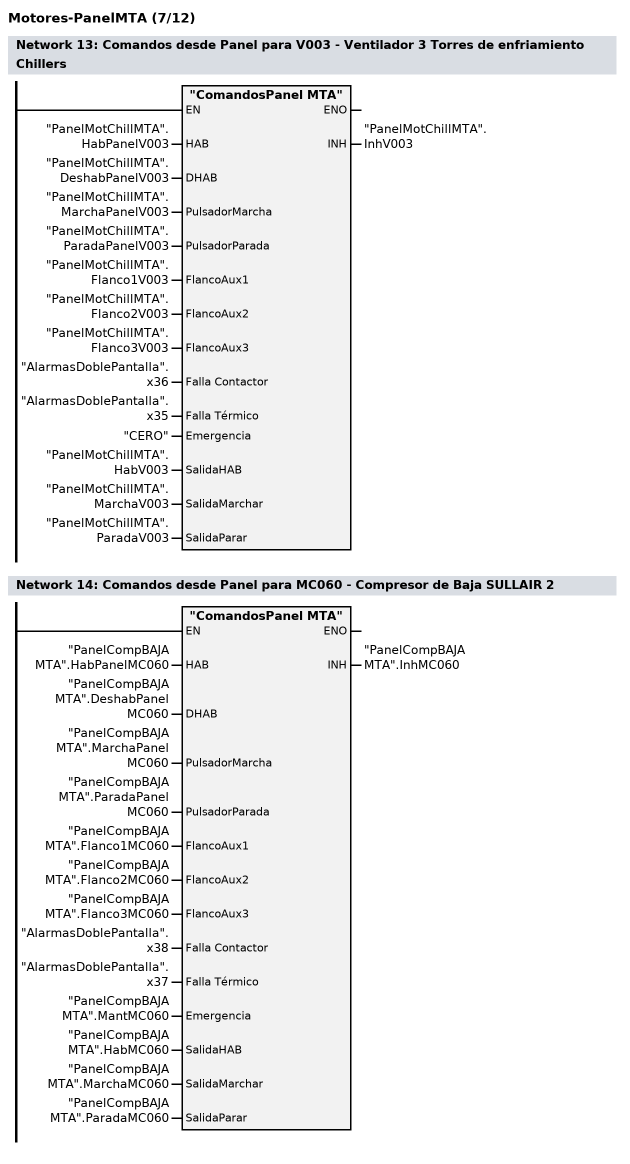
   RUNG wire#powerrail
      "ComandosPanel MTA"(HAB := "PanelMotChillMTA".HabPanelV003, DHAB := "PanelMotChillMTA".DeshabPanelV003, PulsadorMarcha := "PanelMotChillMTA".MarchaPanelV003, PulsadorParada := "PanelMotChillMTA".ParadaPanelV003, FlancoAux1 := "PanelMotChillMTA".Flanco1V003, FlancoAux2 := "PanelMotChillMTA".Flanco2V003, FlancoAux3 := "PanelMotChillMTA".Flanco3V003, "Falla Contactor" := "AlarmasDoblePantalla".x36, "Falla Térmico" := "AlarmasDoblePantalla".x35, Emergencia := "CERO", SalidaHAB := "PanelMotChillMTA".HabV003, SalidaMarchar := "PanelMotChillMTA".MarchaV003, SalidaParar := "PanelMotChillMTA".ParadaV003, INH => "PanelMotChillMTA".InhV003)
   END_RUNG
   // the same network as SCL:
   "ComandosPanel MTA"(HAB := "PanelMotChillMTA".HabPanelV003,
                       DHAB := "PanelMotChillMTA".DeshabPanelV003,
                       PulsadorMarcha := "PanelMotChillMTA".MarchaPanelV003,
                       PulsadorParada := "PanelMotChillMTA".ParadaPanelV003,
                       FlancoAux1 := "PanelMotChillMTA".Flanco1V003,
                       FlancoAux2 := "PanelMotChillMTA".Flanco2V003,
                       FlancoAux3 := "PanelMotChillMTA".Flanco3V003,
                       "Falla Contactor" := "AlarmasDoblePantalla".x36,
                       "Falla Térmico" := "AlarmasDoblePantalla".x35,
                       Emergencia := "CERO",
                       SalidaHAB := "PanelMotChillMTA".HabV003,
                       SalidaMarchar := "PanelMotChillMTA".MarchaV003,
                       SalidaParar := "PanelMotChillMTA".ParadaV003,
                       INH => "PanelMotChillMTA".InhV003);
END_REGION

REGION Network 14: Comandos desde Panel para MC060 - Compresor de Baja SULLAIR 2
   RUNG wire#powerrail
      "ComandosPanel MTA"(HAB := "PanelCompBAJA MTA".HabPanelMC060, DHAB := "PanelCompBAJA MTA".DeshabPanelMC060, PulsadorMarcha := "PanelCompBAJA MTA".MarchaPanelMC060, PulsadorParada := "PanelCompBAJA MTA".ParadaPanelMC060, FlancoAux1 := "PanelCompBAJA MTA".Flanco1MC060, FlancoAux2 := "PanelCompBAJA MTA".Flanco2MC060, FlancoAux3 := "PanelCompBAJA MTA".Flanco3MC060, "Falla Contactor" := "AlarmasDoblePantalla".x38, "Falla Térmico" := "AlarmasDoblePantalla".x37, Emergencia := "PanelCompBAJA MTA".MantMC060, INH => "PanelCompBAJA MTA".InhMC060, SalidaHAB := "PanelCompBAJA MTA".HabMC060, SalidaMarchar := "PanelCompBAJA MTA".MarchaMC060, SalidaParar := "PanelCompBAJA MTA".ParadaMC060)
   END_RUNG
   // the same network as SCL:
   "ComandosPanel MTA"(HAB := "PanelCompBAJA MTA".HabPanelMC060,
                       DHAB := "PanelCompBAJA MTA".DeshabPanelMC060,
                       PulsadorMarcha := "PanelCompBAJA MTA".MarchaPanelMC060,
                       PulsadorParada := "PanelCompBAJA MTA".ParadaPanelMC060,
                       FlancoAux1 := "PanelCompBAJA MTA".Flanco1MC060,
                       FlancoAux2 := "PanelCompBAJA MTA".Flanco2MC060,
                       FlancoAux3 := "PanelCompBAJA MTA".Flanco3MC060,
                       "Falla Contactor" := "AlarmasDoblePantalla".x38,
                       "Falla Térmico" := "AlarmasDoblePantalla".x37,
                       Emergencia := "PanelCompBAJA MTA".MantMC060,
                       SalidaHAB := "PanelCompBAJA MTA".HabMC060,
                       SalidaMarchar := "PanelCompBAJA MTA".MarchaMC060,
                       SalidaParar := "PanelCompBAJA MTA".ParadaMC060,
                       INH => "PanelCompBAJA MTA".InhMC060);
END_REGION

REGION Network 15: Comandos desde Panel para MC061 - Compresor de Baja SULLAIR 1
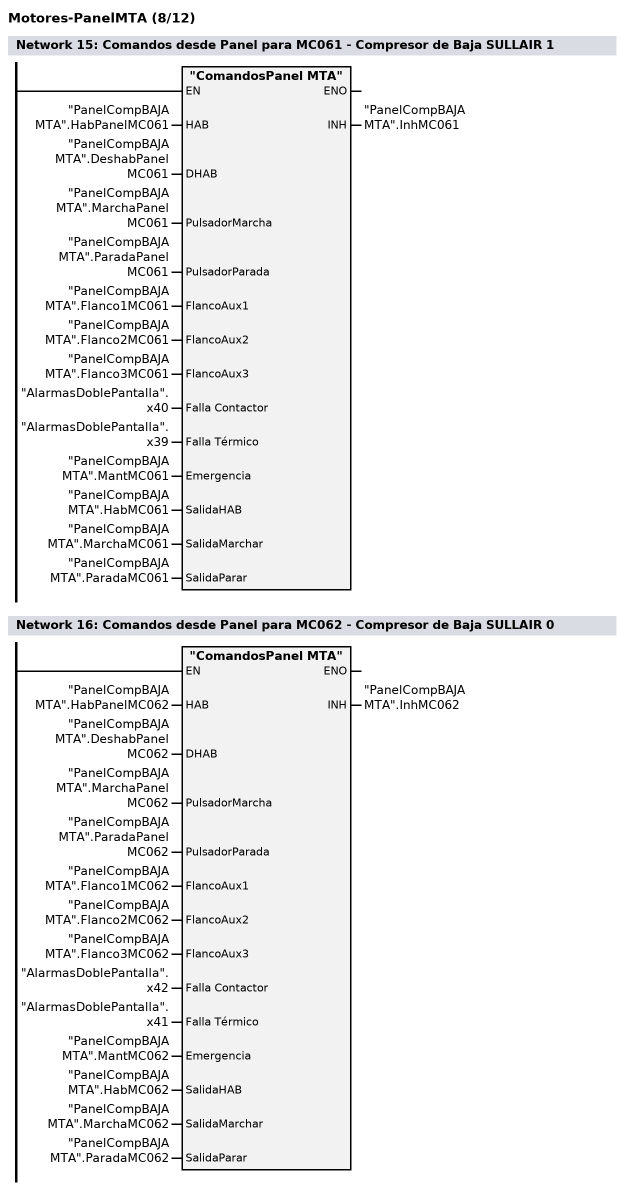
   RUNG wire#powerrail
      "ComandosPanel MTA"(HAB := "PanelCompBAJA MTA".HabPanelMC061, DHAB := "PanelCompBAJA MTA".DeshabPanelMC061, PulsadorMarcha := "PanelCompBAJA MTA".MarchaPanelMC061, PulsadorParada := "PanelCompBAJA MTA".ParadaPanelMC061, FlancoAux1 := "PanelCompBAJA MTA".Flanco1MC061, FlancoAux2 := "PanelCompBAJA MTA".Flanco2MC061, FlancoAux3 := "PanelCompBAJA MTA".Flanco3MC061, "Falla Contactor" := "AlarmasDoblePantalla".x40, "Falla Térmico" := "AlarmasDoblePantalla".x39, Emergencia := "PanelCompBAJA MTA".MantMC061, INH => "PanelCompBAJA MTA".InhMC061, SalidaHAB := "PanelCompBAJA MTA".HabMC061, SalidaMarchar := "PanelCompBAJA MTA".MarchaMC061, SalidaParar := "PanelCompBAJA MTA".ParadaMC061)
   END_RUNG
   // the same network as SCL:
   "ComandosPanel MTA"(HAB := "PanelCompBAJA MTA".HabPanelMC061,
                       DHAB := "PanelCompBAJA MTA".DeshabPanelMC061,
                       PulsadorMarcha := "PanelCompBAJA MTA".MarchaPanelMC061,
                       PulsadorParada := "PanelCompBAJA MTA".ParadaPanelMC061,
                       FlancoAux1 := "PanelCompBAJA MTA".Flanco1MC061,
                       FlancoAux2 := "PanelCompBAJA MTA".Flanco2MC061,
                       FlancoAux3 := "PanelCompBAJA MTA".Flanco3MC061,
                       "Falla Contactor" := "AlarmasDoblePantalla".x40,
                       "Falla Térmico" := "AlarmasDoblePantalla".x39,
                       Emergencia := "PanelCompBAJA MTA".MantMC061,
                       SalidaHAB := "PanelCompBAJA MTA".HabMC061,
                       SalidaMarchar := "PanelCompBAJA MTA".MarchaMC061,
                       SalidaParar := "PanelCompBAJA MTA".ParadaMC061,
                       INH => "PanelCompBAJA MTA".InhMC061);
END_REGION

REGION Network 16: Comandos desde Panel para MC062 - Compresor de Baja SULLAIR 0
   RUNG wire#powerrail
      "ComandosPanel MTA"(HAB := "PanelCompBAJA MTA".HabPanelMC062, DHAB := "PanelCompBAJA MTA".DeshabPanelMC062, PulsadorMarcha := "PanelCompBAJA MTA".MarchaPanelMC062, PulsadorParada := "PanelCompBAJA MTA".ParadaPanelMC062, FlancoAux1 := "PanelCompBAJA MTA".Flanco1MC062, FlancoAux2 := "PanelCompBAJA MTA".Flanco2MC062, FlancoAux3 := "PanelCompBAJA MTA".Flanco3MC062, "Falla Contactor" := "AlarmasDoblePantalla".x42, "Falla Térmico" := "AlarmasDoblePantalla".x41, Emergencia := "PanelCompBAJA MTA".MantMC062, INH => "PanelCompBAJA MTA".InhMC062, SalidaHAB := "PanelCompBAJA MTA".HabMC062, SalidaMarchar := "PanelCompBAJA MTA".MarchaMC062, SalidaParar := "PanelCompBAJA MTA".ParadaMC062)
   END_RUNG
   // the same network as SCL:
   "ComandosPanel MTA"(HAB := "PanelCompBAJA MTA".HabPanelMC062,
                       DHAB := "PanelCompBAJA MTA".DeshabPanelMC062,
                       PulsadorMarcha := "PanelCompBAJA MTA".MarchaPanelMC062,
                       PulsadorParada := "PanelCompBAJA MTA".ParadaPanelMC062,
                       FlancoAux1 := "PanelCompBAJA MTA".Flanco1MC062,
                       FlancoAux2 := "PanelCompBAJA MTA".Flanco2MC062,
                       FlancoAux3 := "PanelCompBAJA MTA".Flanco3MC062,
                       "Falla Contactor" := "AlarmasDoblePantalla".x42,
                       "Falla Térmico" := "AlarmasDoblePantalla".x41,
                       Emergencia := "PanelCompBAJA MTA".MantMC062,
                       SalidaHAB := "PanelCompBAJA MTA".HabMC062,
                       SalidaMarchar := "PanelCompBAJA MTA".MarchaMC062,
                       SalidaParar := "PanelCompBAJA MTA".ParadaMC062,
                       INH => "PanelCompBAJA MTA".InhMC062);
END_REGION

REGION Network 17: Comandos desde Panel para MC063 - Compresor de Baja ATLAS 3
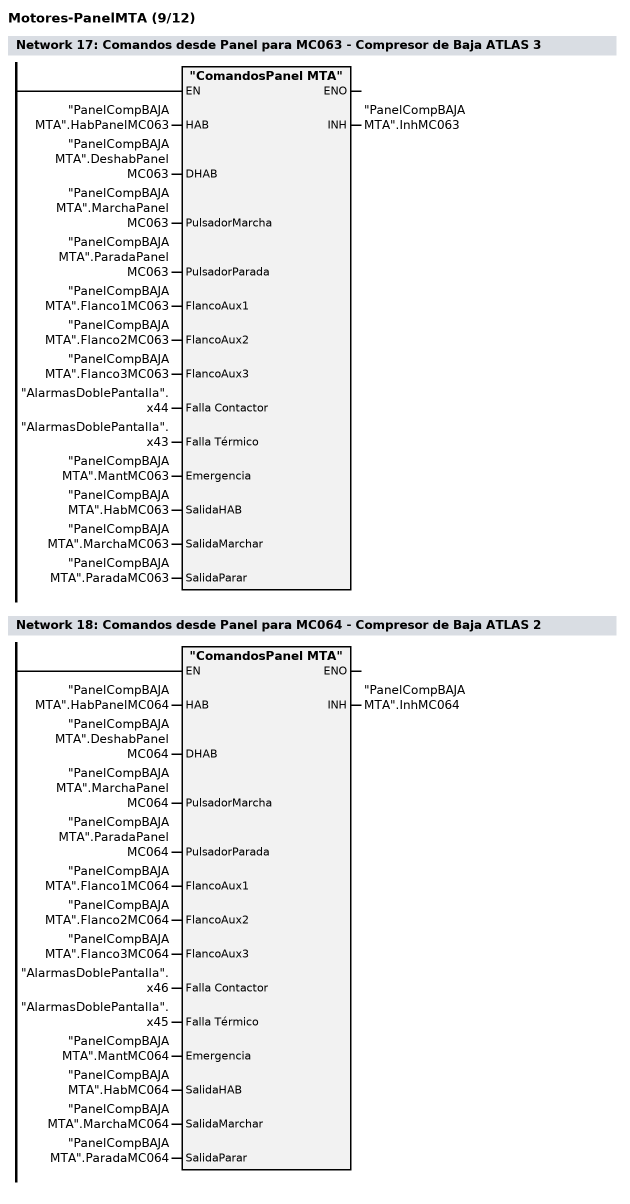
   RUNG wire#powerrail
      "ComandosPanel MTA"(HAB := "PanelCompBAJA MTA".HabPanelMC063, DHAB := "PanelCompBAJA MTA".DeshabPanelMC063, PulsadorMarcha := "PanelCompBAJA MTA".MarchaPanelMC063, PulsadorParada := "PanelCompBAJA MTA".ParadaPanelMC063, FlancoAux1 := "PanelCompBAJA MTA".Flanco1MC063, FlancoAux2 := "PanelCompBAJA MTA".Flanco2MC063, FlancoAux3 := "PanelCompBAJA MTA".Flanco3MC063, "Falla Contactor" := "AlarmasDoblePantalla".x44, "Falla Térmico" := "AlarmasDoblePantalla".x43, Emergencia := "PanelCompBAJA MTA".MantMC063, INH => "PanelCompBAJA MTA".InhMC063, SalidaHAB := "PanelCompBAJA MTA".HabMC063, SalidaMarchar := "PanelCompBAJA MTA".MarchaMC063, SalidaParar := "PanelCompBAJA MTA".ParadaMC063)
   END_RUNG
   // the same network as SCL:
   "ComandosPanel MTA"(HAB := "PanelCompBAJA MTA".HabPanelMC063,
                       DHAB := "PanelCompBAJA MTA".DeshabPanelMC063,
                       PulsadorMarcha := "PanelCompBAJA MTA".MarchaPanelMC063,
                       PulsadorParada := "PanelCompBAJA MTA".ParadaPanelMC063,
                       FlancoAux1 := "PanelCompBAJA MTA".Flanco1MC063,
                       FlancoAux2 := "PanelCompBAJA MTA".Flanco2MC063,
                       FlancoAux3 := "PanelCompBAJA MTA".Flanco3MC063,
                       "Falla Contactor" := "AlarmasDoblePantalla".x44,
                       "Falla Térmico" := "AlarmasDoblePantalla".x43,
                       Emergencia := "PanelCompBAJA MTA".MantMC063,
                       SalidaHAB := "PanelCompBAJA MTA".HabMC063,
                       SalidaMarchar := "PanelCompBAJA MTA".MarchaMC063,
                       SalidaParar := "PanelCompBAJA MTA".ParadaMC063,
                       INH => "PanelCompBAJA MTA".InhMC063);
END_REGION

REGION Network 18: Comandos desde Panel para MC064 - Compresor de Baja ATLAS 2
   RUNG wire#powerrail
      "ComandosPanel MTA"(HAB := "PanelCompBAJA MTA".HabPanelMC064, DHAB := "PanelCompBAJA MTA".DeshabPanelMC064, PulsadorMarcha := "PanelCompBAJA MTA".MarchaPanelMC064, PulsadorParada := "PanelCompBAJA MTA".ParadaPanelMC064, FlancoAux1 := "PanelCompBAJA MTA".Flanco1MC064, FlancoAux2 := "PanelCompBAJA MTA".Flanco2MC064, FlancoAux3 := "PanelCompBAJA MTA".Flanco3MC064, "Falla Contactor" := "AlarmasDoblePantalla".x46, "Falla Térmico" := "AlarmasDoblePantalla".x45, Emergencia := "PanelCompBAJA MTA".MantMC064, INH => "PanelCompBAJA MTA".InhMC064, SalidaHAB := "PanelCompBAJA MTA".HabMC064, SalidaMarchar := "PanelCompBAJA MTA".MarchaMC064, SalidaParar := "PanelCompBAJA MTA".ParadaMC064)
   END_RUNG
   // the same network as SCL:
   "ComandosPanel MTA"(HAB := "PanelCompBAJA MTA".HabPanelMC064,
                       DHAB := "PanelCompBAJA MTA".DeshabPanelMC064,
                       PulsadorMarcha := "PanelCompBAJA MTA".MarchaPanelMC064,
                       PulsadorParada := "PanelCompBAJA MTA".ParadaPanelMC064,
                       FlancoAux1 := "PanelCompBAJA MTA".Flanco1MC064,
                       FlancoAux2 := "PanelCompBAJA MTA".Flanco2MC064,
                       FlancoAux3 := "PanelCompBAJA MTA".Flanco3MC064,
                       "Falla Contactor" := "AlarmasDoblePantalla".x46,
                       "Falla Térmico" := "AlarmasDoblePantalla".x45,
                       Emergencia := "PanelCompBAJA MTA".MantMC064,
                       SalidaHAB := "PanelCompBAJA MTA".HabMC064,
                       SalidaMarchar := "PanelCompBAJA MTA".MarchaMC064,
                       SalidaParar := "PanelCompBAJA MTA".ParadaMC064,
                       INH => "PanelCompBAJA MTA".InhMC064);
END_REGION

REGION Network 19: Comandos desde Panel para MS050 - Secador de Alta ABC1
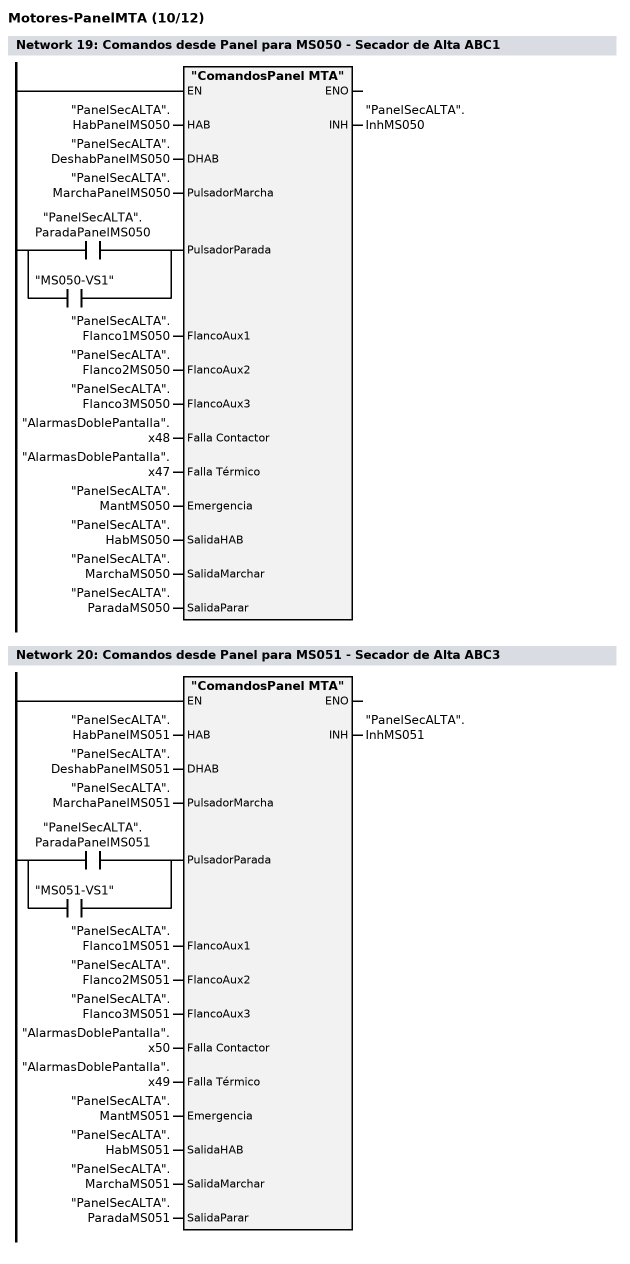
   RUNG wire#powerrail
      "ComandosPanel MTA"(HAB := "PanelSecALTA".HabPanelMS050, DHAB := "PanelSecALTA".DeshabPanelMS050, PulsadorMarcha := "PanelSecALTA".MarchaPanelMS050, PulsadorParada := wire#w1, FlancoAux1 := "PanelSecALTA".Flanco1MS050, FlancoAux2 := "PanelSecALTA".Flanco2MS050, FlancoAux3 := "PanelSecALTA".Flanco3MS050, "Falla Contactor" := "AlarmasDoblePantalla".x48, "Falla Térmico" := "AlarmasDoblePantalla".x47, Emergencia := "PanelSecALTA".MantMS050, INH => "PanelSecALTA".InhMS050, SalidaHAB := "PanelSecALTA".HabMS050, SalidaMarchar := "PanelSecALTA".MarchaMS050, SalidaParar := "PanelSecALTA".ParadaMS050)
   END_RUNG
   RUNG wire#powerrail
      Contact( "PanelSecALTA".ParadaPanelMS050 )
   END_RUNG wire#w1
   RUNG wire#powerrail
      Contact( "MS050-VS1" )
   END_RUNG wire#w1
   // the same network as SCL:
   "ComandosPanel MTA"(HAB := "PanelSecALTA".HabPanelMS050,
                       DHAB := "PanelSecALTA".DeshabPanelMS050,
                       PulsadorMarcha := "PanelSecALTA".MarchaPanelMS050,
                       PulsadorParada := "PanelSecALTA".ParadaPanelMS050 OR "MS050-VS1",
                       FlancoAux1 := "PanelSecALTA".Flanco1MS050,
                       FlancoAux2 := "PanelSecALTA".Flanco2MS050,
                       FlancoAux3 := "PanelSecALTA".Flanco3MS050,
                       "Falla Contactor" := "AlarmasDoblePantalla".x48,
                       "Falla Térmico" := "AlarmasDoblePantalla".x47,
                       Emergencia := "PanelSecALTA".MantMS050,
                       SalidaHAB := "PanelSecALTA".HabMS050,
                       SalidaMarchar := "PanelSecALTA".MarchaMS050,
                       SalidaParar := "PanelSecALTA".ParadaMS050,
                       INH => "PanelSecALTA".InhMS050);
END_REGION

REGION Network 20: Comandos desde Panel para MS051 - Secador de Alta ABC3
   RUNG wire#powerrail
      "ComandosPanel MTA"(HAB := "PanelSecALTA".HabPanelMS051, DHAB := "PanelSecALTA".DeshabPanelMS051, PulsadorMarcha := "PanelSecALTA".MarchaPanelMS051, PulsadorParada := wire#w1, FlancoAux1 := "PanelSecALTA".Flanco1MS051, FlancoAux2 := "PanelSecALTA".Flanco2MS051, FlancoAux3 := "PanelSecALTA".Flanco3MS051, "Falla Contactor" := "AlarmasDoblePantalla".x50, "Falla Térmico" := "AlarmasDoblePantalla".x49, Emergencia := "PanelSecALTA".MantMS051, INH => "PanelSecALTA".InhMS051, SalidaHAB := "PanelSecALTA".HabMS051, SalidaMarchar := "PanelSecALTA".MarchaMS051, SalidaParar := "PanelSecALTA".ParadaMS051)
   END_RUNG
   RUNG wire#powerrail
      Contact( "PanelSecALTA".ParadaPanelMS051 )
   END_RUNG wire#w1
   RUNG wire#powerrail
      Contact( "MS051-VS1" )
   END_RUNG wire#w1
   // the same network as SCL:
   "ComandosPanel MTA"(HAB := "PanelSecALTA".HabPanelMS051,
                       DHAB := "PanelSecALTA".DeshabPanelMS051,
                       PulsadorMarcha := "PanelSecALTA".MarchaPanelMS051,
                       PulsadorParada := "PanelSecALTA".ParadaPanelMS051 OR "MS051-VS1",
                       FlancoAux1 := "PanelSecALTA".Flanco1MS051,
                       FlancoAux2 := "PanelSecALTA".Flanco2MS051,
                       FlancoAux3 := "PanelSecALTA".Flanco3MS051,
                       "Falla Contactor" := "AlarmasDoblePantalla".x50,
                       "Falla Térmico" := "AlarmasDoblePantalla".x49,
                       Emergencia := "PanelSecALTA".MantMS051,
                       SalidaHAB := "PanelSecALTA".HabMS051,
                       SalidaMarchar := "PanelSecALTA".MarchaMS051,
                       SalidaParar := "PanelSecALTA".ParadaMS051,
                       INH => "PanelSecALTA".InhMS051);
END_REGION

REGION Network 21: Comandos desde Panel para MS052 - Secador de Alta ABC2
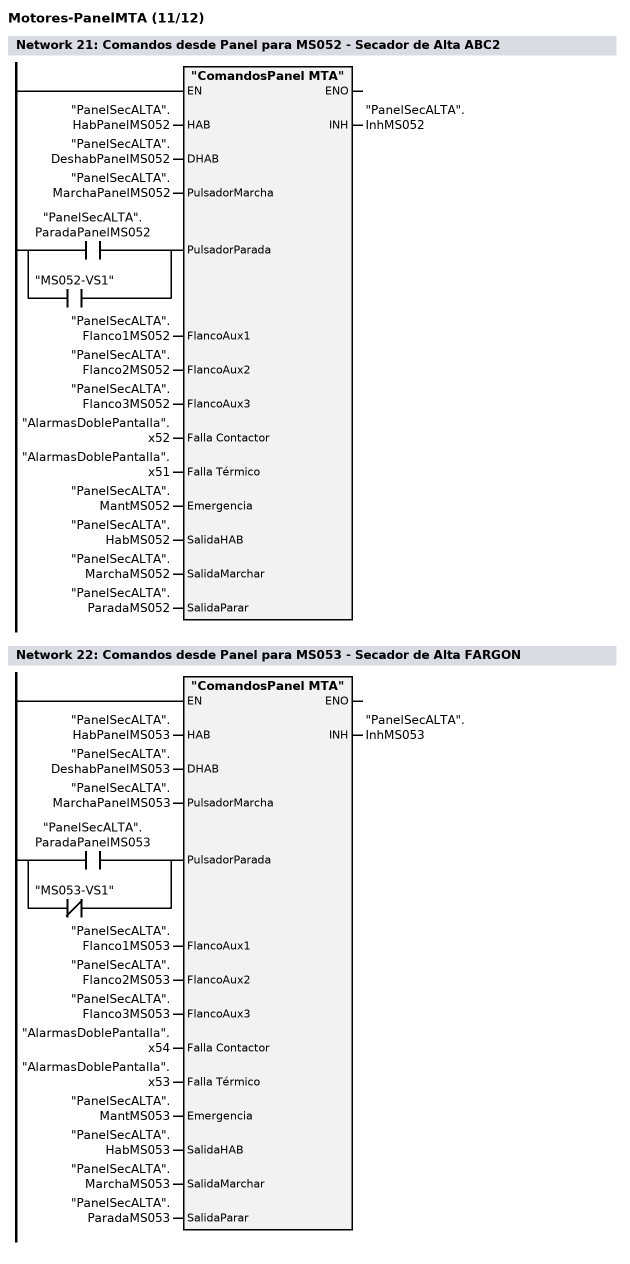
   RUNG wire#powerrail
      "ComandosPanel MTA"(HAB := "PanelSecALTA".HabPanelMS052, DHAB := "PanelSecALTA".DeshabPanelMS052, PulsadorMarcha := "PanelSecALTA".MarchaPanelMS052, PulsadorParada := wire#w1, FlancoAux1 := "PanelSecALTA".Flanco1MS052, FlancoAux2 := "PanelSecALTA".Flanco2MS052, FlancoAux3 := "PanelSecALTA".Flanco3MS052, "Falla Contactor" := "AlarmasDoblePantalla".x52, "Falla Térmico" := "AlarmasDoblePantalla".x51, Emergencia := "PanelSecALTA".MantMS052, INH => "PanelSecALTA".InhMS052, SalidaHAB := "PanelSecALTA".HabMS052, SalidaMarchar := "PanelSecALTA".MarchaMS052, SalidaParar := "PanelSecALTA".ParadaMS052)
   END_RUNG
   RUNG wire#powerrail
      Contact( "PanelSecALTA".ParadaPanelMS052 )
   END_RUNG wire#w1
   RUNG wire#powerrail
      Contact( "MS052-VS1" )
   END_RUNG wire#w1
   // the same network as SCL:
   "ComandosPanel MTA"(HAB := "PanelSecALTA".HabPanelMS052,
                       DHAB := "PanelSecALTA".DeshabPanelMS052,
                       PulsadorMarcha := "PanelSecALTA".MarchaPanelMS052,
                       PulsadorParada := "PanelSecALTA".ParadaPanelMS052 OR "MS052-VS1",
                       FlancoAux1 := "PanelSecALTA".Flanco1MS052,
                       FlancoAux2 := "PanelSecALTA".Flanco2MS052,
                       FlancoAux3 := "PanelSecALTA".Flanco3MS052,
                       "Falla Contactor" := "AlarmasDoblePantalla".x52,
                       "Falla Térmico" := "AlarmasDoblePantalla".x51,
                       Emergencia := "PanelSecALTA".MantMS052,
                       SalidaHAB := "PanelSecALTA".HabMS052,
                       SalidaMarchar := "PanelSecALTA".MarchaMS052,
                       SalidaParar := "PanelSecALTA".ParadaMS052,
                       INH => "PanelSecALTA".InhMS052);
END_REGION

REGION Network 22: Comandos desde Panel para MS053 - Secador de Alta FARGON
   RUNG wire#powerrail
      "ComandosPanel MTA"(HAB := "PanelSecALTA".HabPanelMS053, DHAB := "PanelSecALTA".DeshabPanelMS053, PulsadorMarcha := "PanelSecALTA".MarchaPanelMS053, PulsadorParada := wire#w1, FlancoAux1 := "PanelSecALTA".Flanco1MS053, FlancoAux2 := "PanelSecALTA".Flanco2MS053, FlancoAux3 := "PanelSecALTA".Flanco3MS053, "Falla Contactor" := "AlarmasDoblePantalla".x54, "Falla Térmico" := "AlarmasDoblePantalla".x53, Emergencia := "PanelSecALTA".MantMS053, INH => "PanelSecALTA".InhMS053, SalidaHAB := "PanelSecALTA".HabMS053, SalidaMarchar := "PanelSecALTA".MarchaMS053, SalidaParar := "PanelSecALTA".ParadaMS053)
   END_RUNG
   RUNG wire#powerrail
      Contact( "PanelSecALTA".ParadaPanelMS053 )
   END_RUNG wire#w1
   RUNG wire#powerrail
      I_Contact( "MS053-VS1" )
   END_RUNG wire#w1
   // the same network as SCL:
   "ComandosPanel MTA"(HAB := "PanelSecALTA".HabPanelMS053,
                       DHAB := "PanelSecALTA".DeshabPanelMS053,
                       PulsadorMarcha := "PanelSecALTA".MarchaPanelMS053,
                       PulsadorParada := "PanelSecALTA".ParadaPanelMS053 OR NOT "MS053-VS1",
                       FlancoAux1 := "PanelSecALTA".Flanco1MS053,
                       FlancoAux2 := "PanelSecALTA".Flanco2MS053,
                       FlancoAux3 := "PanelSecALTA".Flanco3MS053,
                       "Falla Contactor" := "AlarmasDoblePantalla".x54,
                       "Falla Térmico" := "AlarmasDoblePantalla".x53,
                       Emergencia := "PanelSecALTA".MantMS053,
                       SalidaHAB := "PanelSecALTA".HabMS053,
                       SalidaMarchar := "PanelSecALTA".MarchaMS053,
                       SalidaParar := "PanelSecALTA".ParadaMS053,
                       INH => "PanelSecALTA".InhMS053);
END_REGION

REGION Network 23: Comandos desde Panel para MS054 - Secador de Baja SULLAIR 1
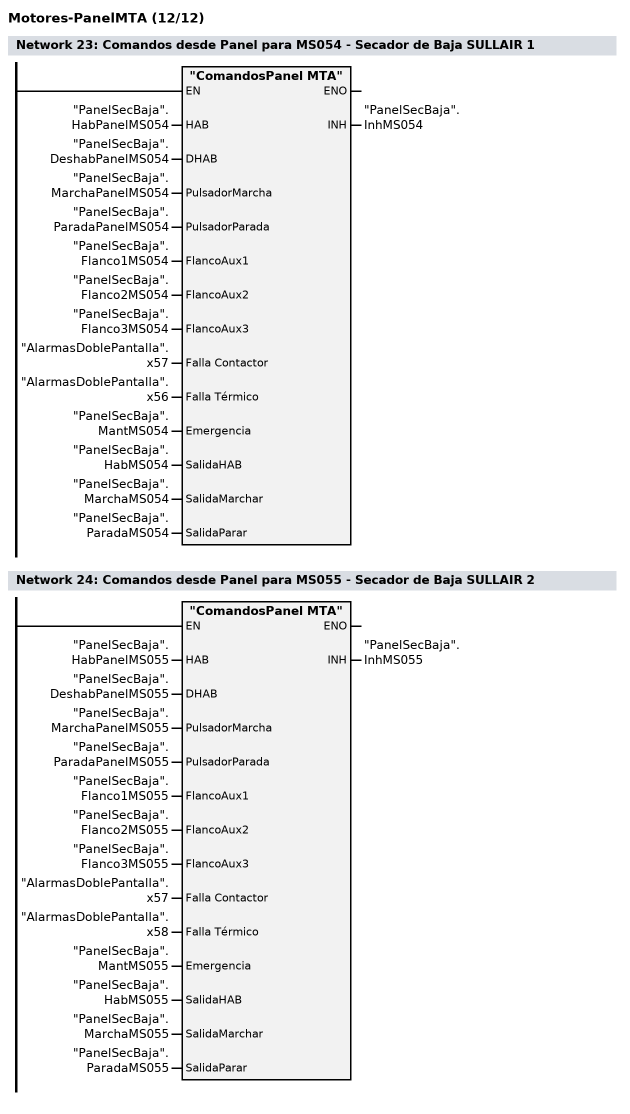
   RUNG wire#powerrail
      "ComandosPanel MTA"(HAB := "PanelSecBaja".HabPanelMS054, DHAB := "PanelSecBaja".DeshabPanelMS054, PulsadorMarcha := "PanelSecBaja".MarchaPanelMS054, PulsadorParada := "PanelSecBaja".ParadaPanelMS054, FlancoAux1 := "PanelSecBaja".Flanco1MS054, FlancoAux2 := "PanelSecBaja".Flanco2MS054, FlancoAux3 := "PanelSecBaja".Flanco3MS054, "Falla Contactor" := "AlarmasDoblePantalla".x57, "Falla Térmico" := "AlarmasDoblePantalla".x56, Emergencia := "PanelSecBaja".MantMS054, INH => "PanelSecBaja".InhMS054, SalidaHAB := "PanelSecBaja".HabMS054, SalidaMarchar := "PanelSecBaja".MarchaMS054, SalidaParar := "PanelSecBaja".ParadaMS054)
   END_RUNG
   // the same network as SCL:
   "ComandosPanel MTA"(HAB := "PanelSecBaja".HabPanelMS054,
                       DHAB := "PanelSecBaja".DeshabPanelMS054,
                       PulsadorMarcha := "PanelSecBaja".MarchaPanelMS054,
                       PulsadorParada := "PanelSecBaja".ParadaPanelMS054,
                       FlancoAux1 := "PanelSecBaja".Flanco1MS054,
                       FlancoAux2 := "PanelSecBaja".Flanco2MS054,
                       FlancoAux3 := "PanelSecBaja".Flanco3MS054,
                       "Falla Contactor" := "AlarmasDoblePantalla".x57,
                       "Falla Térmico" := "AlarmasDoblePantalla".x56,
                       Emergencia := "PanelSecBaja".MantMS054,
                       SalidaHAB := "PanelSecBaja".HabMS054,
                       SalidaMarchar := "PanelSecBaja".MarchaMS054,
                       SalidaParar := "PanelSecBaja".ParadaMS054,
                       INH => "PanelSecBaja".InhMS054);
END_REGION

REGION Network 24: Comandos desde Panel para MS055 - Secador de Baja SULLAIR 2
   RUNG wire#powerrail
      "ComandosPanel MTA"(HAB := "PanelSecBaja".HabPanelMS055, DHAB := "PanelSecBaja".DeshabPanelMS055, PulsadorMarcha := "PanelSecBaja".MarchaPanelMS055, PulsadorParada := "PanelSecBaja".ParadaPanelMS055, FlancoAux1 := "PanelSecBaja".Flanco1MS055, FlancoAux2 := "PanelSecBaja".Flanco2MS055, FlancoAux3 := "PanelSecBaja".Flanco3MS055, "Falla Contactor" := "AlarmasDoblePantalla".x57, "Falla Térmico" := "AlarmasDoblePantalla".x58, Emergencia := "PanelSecBaja".MantMS055, INH => "PanelSecBaja".InhMS055, SalidaHAB := "PanelSecBaja".HabMS055, SalidaMarchar := "PanelSecBaja".MarchaMS055, SalidaParar := "PanelSecBaja".ParadaMS055)
   END_RUNG
   // the same network as SCL:
   "ComandosPanel MTA"(HAB := "PanelSecBaja".HabPanelMS055,
                       DHAB := "PanelSecBaja".DeshabPanelMS055,
                       PulsadorMarcha := "PanelSecBaja".MarchaPanelMS055,
                       PulsadorParada := "PanelSecBaja".ParadaPanelMS055,
                       FlancoAux1 := "PanelSecBaja".Flanco1MS055,
                       FlancoAux2 := "PanelSecBaja".Flanco2MS055,
                       FlancoAux3 := "PanelSecBaja".Flanco3MS055,
                       "Falla Contactor" := "AlarmasDoblePantalla".x57,
                       "Falla Térmico" := "AlarmasDoblePantalla".x58,
                       Emergencia := "PanelSecBaja".MantMS055,
                       SalidaHAB := "PanelSecBaja".HabMS055,
                       SalidaMarchar := "PanelSecBaja".MarchaMS055,
                       SalidaParar := "PanelSecBaja".ParadaMS055,
                       INH => "PanelSecBaja".InhMS055);
END_REGION
END_FUNCTION

FUNCTION "ComandosPanel MTA" : Void   // FC19, LAD
{ S7_Optimized_Access := 'FALSE' }
VERSION : 0.1
   VAR_INPUT
      HAB : Bool;   // Habilitación
      DHAB : Bool;   // Deshabilitación
      PulsadorMarcha : Bool;   // Pulsador de Marcha
      PulsadorParada : Bool;   // Pulsador de Parada
      FlancoAux1 : Bool;
      FlancoAux2 : Bool;
      FlancoAux3 : Bool;
      "Falla Contactor" : Bool;   // Falla Contactor
      "Falla Térmico" : Bool;   // Falla Térmico
      Emergencia : Bool;
   END_VAR
   VAR_OUTPUT
      INH : Bool;
   END_VAR
   VAR_IN_OUT
      SalidaHAB : Bool;
      SalidaMarchar : Bool;
      SalidaParar : Bool;
   END_VAR
   VAR_TEMP   // added for the SCL form of the ladder/FBD networks
      _w1 : Bool;
   END_VAR
BEGIN

REGION Network 1
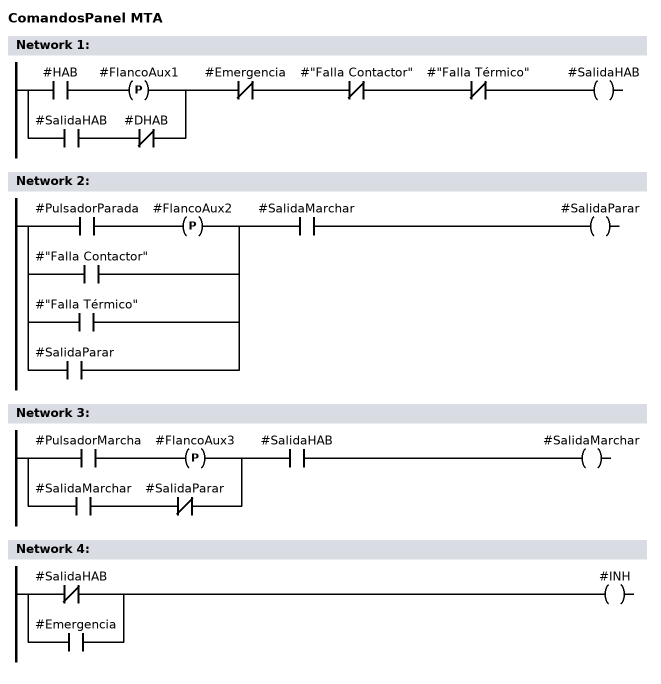
   RUNG wire#powerrail
      Contact( #HAB )
      P_Trig( #FlancoAux1 )
      wire#w1
      I_Contact( #Emergencia )
      I_Contact( #"Falla Contactor" )
      I_Contact( #"Falla Térmico" )
      Coil( #SalidaHAB )
   END_RUNG
   RUNG wire#powerrail
      Contact( #SalidaHAB )
      I_Contact( #DHAB )
   END_RUNG wire#w1
   // the same network as SCL:
   #_w1 := #HAB AND NOT #FlancoAux1;   // rising edge
   #FlancoAux1 := #HAB;
   #SalidaHAB := (#_w1 OR (#SalidaHAB AND NOT #DHAB)) AND NOT #Emergencia AND NOT #"Falla Contactor" AND NOT #"Falla Térmico";
END_REGION

REGION Network 2
   RUNG wire#powerrail
      Contact( #PulsadorParada )
      P_Trig( #FlancoAux2 )
      wire#w1
      Contact( #SalidaMarchar )
      Coil( #SalidaParar )
   END_RUNG
   RUNG wire#powerrail
      Contact( #"Falla Contactor" )
   END_RUNG wire#w1
   RUNG wire#powerrail
      Contact( #"Falla Térmico" )
   END_RUNG wire#w1
   RUNG wire#powerrail
      Contact( #SalidaParar )
   END_RUNG wire#w1
   // the same network as SCL:
   #_w1 := #PulsadorParada AND NOT #FlancoAux2;   // rising edge
   #FlancoAux2 := #PulsadorParada;
   #SalidaParar := (#_w1 OR #"Falla Contactor" OR #"Falla Térmico" OR #SalidaParar) AND #SalidaMarchar;
END_REGION

REGION Network 3
   RUNG wire#powerrail
      Contact( #PulsadorMarcha )
      P_Trig( #FlancoAux3 )
      wire#w1
      Contact( #SalidaHAB )
      Coil( #SalidaMarchar )
   END_RUNG
   RUNG wire#powerrail
      Contact( #SalidaMarchar )
      I_Contact( #SalidaParar )
   END_RUNG wire#w1
   // the same network as SCL:
   #_w1 := #PulsadorMarcha AND NOT #FlancoAux3;   // rising edge
   #FlancoAux3 := #PulsadorMarcha;
   #SalidaMarchar := (#_w1 OR (#SalidaMarchar AND NOT #SalidaParar)) AND #SalidaHAB;
END_REGION

REGION Network 4
   RUNG wire#powerrail
      I_Contact( #SalidaHAB )
      wire#w1
      Coil( #INH )
   END_RUNG
   RUNG wire#powerrail
      Contact( #Emergencia )
   END_RUNG wire#w1
   // the same network as SCL:
   #INH := NOT #SalidaHAB OR #Emergencia;
END_REGION
END_FUNCTION

FUNCTION "FC-ANIM-CMP" : Void   // FC43, LAD
{ S7_Optimized_Access := 'FALSE' }
VERSION : 0.1
   VAR_INPUT
      IN0 : Word;
   END_VAR
   VAR_OUTPUT
      OUT1 : Int;
   END_VAR
BEGIN

REGION Network 1